REGION Network 5: RIO02 4P, 4S Vent A and Vent B control
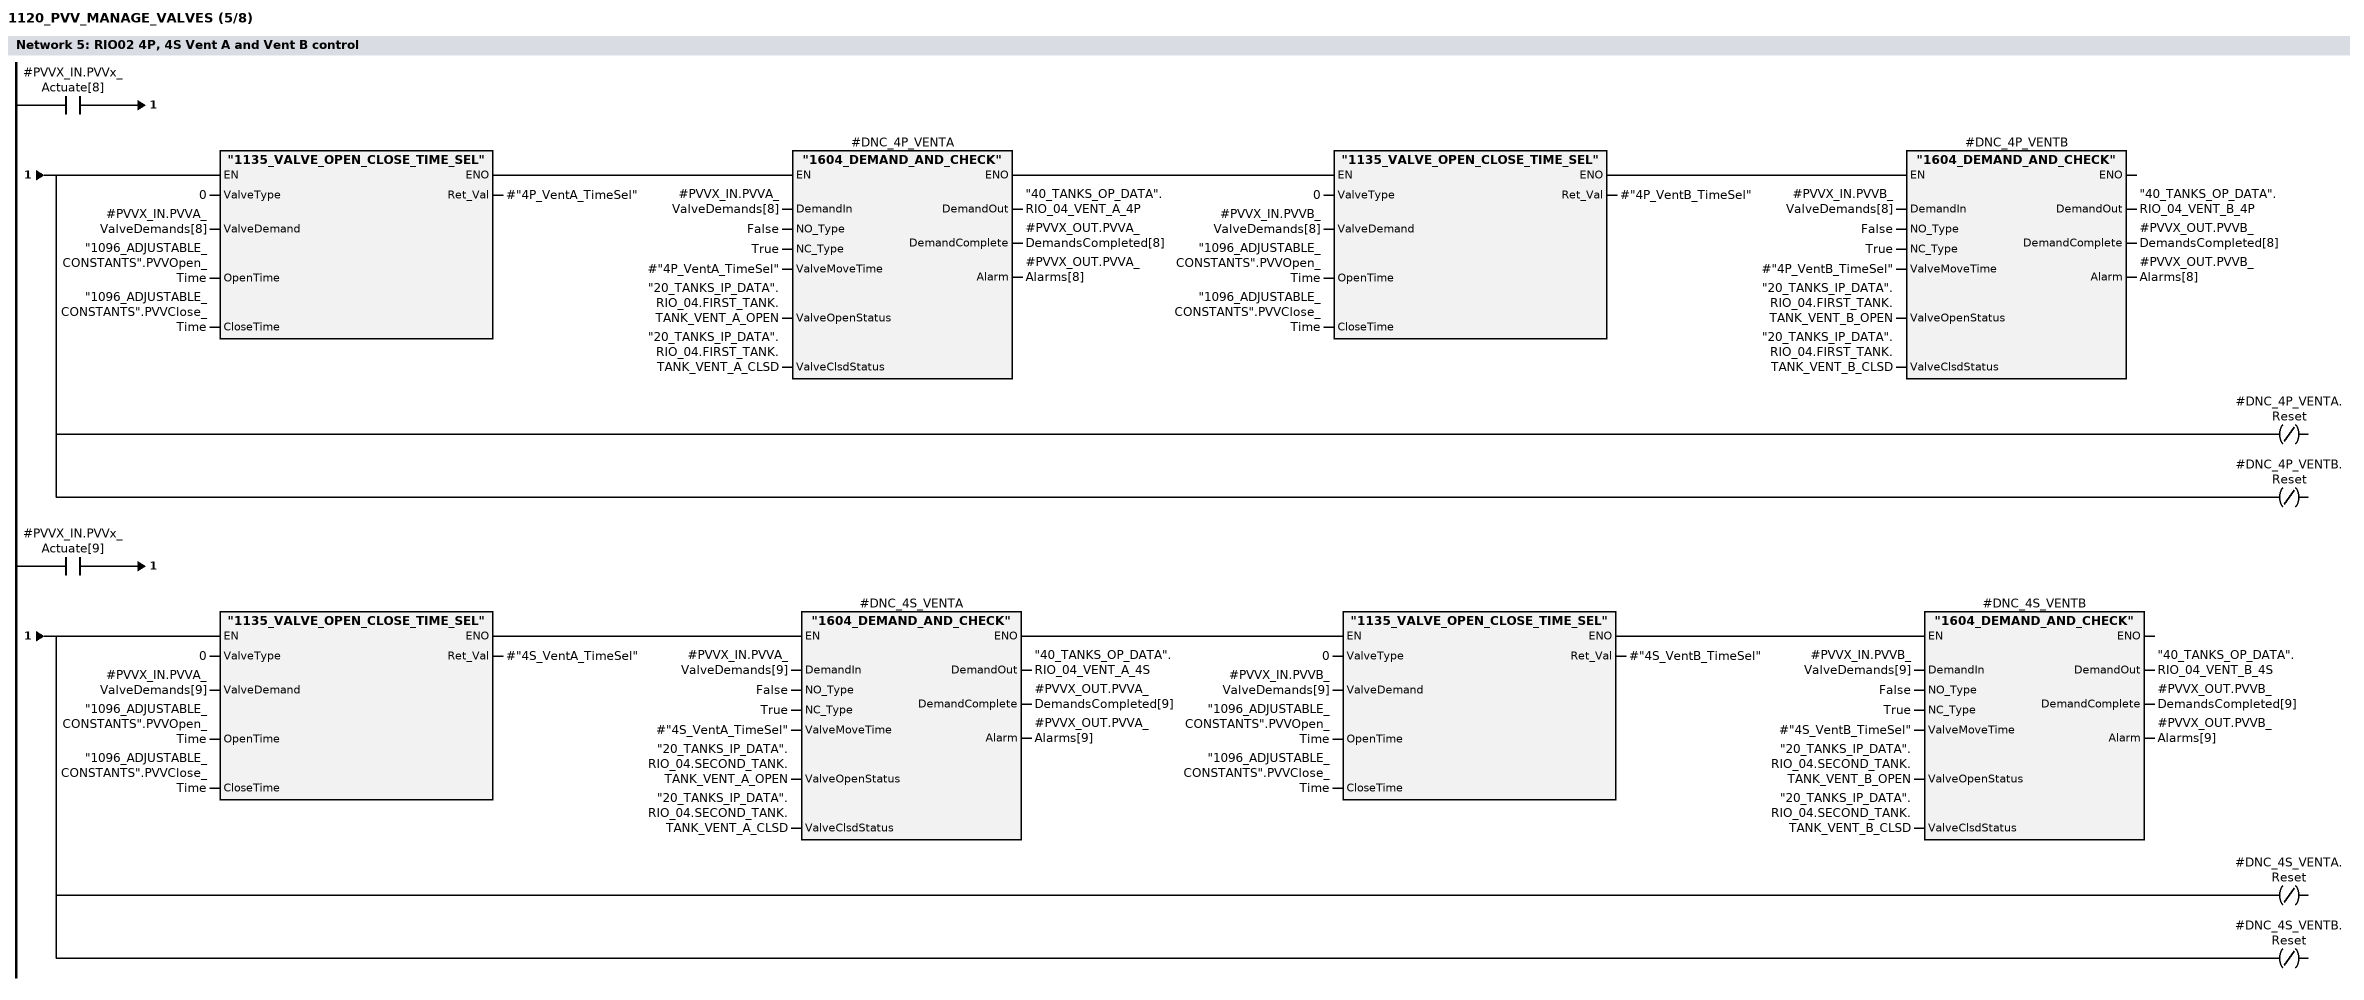
   RUNG wire#powerrail
      Contact( #PVVX_IN.PVVx_Actuate[8] )
      wire#w1
      "1135_VALVE_OPEN_CLOSE_TIME_SEL"(ValveType := 0, ValveDemand := #PVVX_IN.PVVA_ValveDemands[8], OpenTime := "1096_ADJUSTABLE_CONSTANTS".PVVOpen_Time, CloseTime := "1096_ADJUSTABLE_CONSTANTS".PVVClose_Time, Ret_Val => #"4P_VentA_TimeSel")
      #DNC_4P_VENTA(DemandIn := #PVVX_IN.PVVA_ValveDemands[8], NO_Type := False, NC_Type := True, ValveMoveTime := #"4P_VentA_TimeSel", ValveOpenStatus := "20_TANKS_IP_DATA".RIO_04.FIRST_TANK.TANK_VENT_A_OPEN, ValveClsdStatus := "20_TANKS_IP_DATA".RIO_04.FIRST_TANK.TANK_VENT_A_CLSD, DemandOut => "40_TANKS_OP_DATA".RIO_04_VENT_A_4P, DemandComplete => #PVVX_OUT.PVVA_DemandsCompleted[8], Alarm => #PVVX_OUT.PVVA_Alarms[8])
      "1135_VALVE_OPEN_CLOSE_TIME_SEL"(ValveType := 0, ValveDemand := #PVVX_IN.PVVB_ValveDemands[8], OpenTime := "1096_ADJUSTABLE_CONSTANTS".PVVOpen_Time, CloseTime := "1096_ADJUSTABLE_CONSTANTS".PVVClose_Time, Ret_Val => #"4P_VentB_TimeSel")
      #DNC_4P_VENTB(DemandIn := #PVVX_IN.PVVB_ValveDemands[8], NO_Type := False, NC_Type := True, ValveMoveTime := #"4P_VentB_TimeSel", ValveOpenStatus := "20_TANKS_IP_DATA".RIO_04.FIRST_TANK.TANK_VENT_B_OPEN, ValveClsdStatus := "20_TANKS_IP_DATA".RIO_04.FIRST_TANK.TANK_VENT_B_CLSD, DemandOut => "40_TANKS_OP_DATA".RIO_04_VENT_B_4P, DemandComplete => #PVVX_OUT.PVVB_DemandsCompleted[8], Alarm => #PVVX_OUT.PVVB_Alarms[8])
   END_RUNG
   RUNG wire#w1
      I_Coil( #DNC_4P_VENTA.Reset )
   END_RUNG
   RUNG wire#w1
      I_Coil( #DNC_4P_VENTB.Reset )
   END_RUNG
   RUNG wire#powerrail
      Contact( #PVVX_IN.PVVx_Actuate[9] )
      wire#w2
      "1135_VALVE_OPEN_CLOSE_TIME_SEL"(ValveType := 0, ValveDemand := #PVVX_IN.PVVA_ValveDemands[9], OpenTime := "1096_ADJUSTABLE_CONSTANTS".PVVOpen_Time, CloseTime := "1096_ADJUSTABLE_CONSTANTS".PVVClose_Time, Ret_Val => #"4S_VentA_TimeSel")
      #DNC_4S_VENTA(DemandIn := #PVVX_IN.PVVA_ValveDemands[9], NO_Type := False, NC_Type := True, ValveMoveTime := #"4S_VentA_TimeSel", ValveOpenStatus := "20_TANKS_IP_DATA".RIO_04.SECOND_TANK.TANK_VENT_A_OPEN, ValveClsdStatus := "20_TANKS_IP_DATA".RIO_04.SECOND_TANK.TANK_VENT_A_CLSD, DemandOut => "40_TANKS_OP_DATA".RIO_04_VENT_A_4S, DemandComplete => #PVVX_OUT.PVVA_DemandsCompleted[9], Alarm => #PVVX_OUT.PVVA_Alarms[9])
      "1135_VALVE_OPEN_CLOSE_TIME_SEL"(ValveType := 0, ValveDemand := #PVVX_IN.PVVB_ValveDemands[9], OpenTime := "1096_ADJUSTABLE_CONSTANTS".PVVOpen_Time, CloseTime := "1096_ADJUSTABLE_CONSTANTS".PVVClose_Time, Ret_Val => #"4S_VentB_TimeSel")
      #DNC_4S_VENTB(DemandIn := #PVVX_IN.PVVB_ValveDemands[9], NO_Type := False, NC_Type := True, ValveMoveTime := #"4S_VentB_TimeSel", ValveOpenStatus := "20_TANKS_IP_DATA".RIO_04.SECOND_TANK.TANK_VENT_B_OPEN, ValveClsdStatus := "20_TANKS_IP_DATA".RIO_04.SECOND_TANK.TANK_VENT_B_CLSD, DemandOut => "40_TANKS_OP_DATA".RIO_04_VENT_B_4S, DemandComplete => #PVVX_OUT.PVVB_DemandsCompleted[9], Alarm => #PVVX_OUT.PVVB_Alarms[9])
   END_RUNG
   RUNG wire#w2
      I_Coil( #DNC_4S_VENTA.Reset )
   END_RUNG
   RUNG wire#w2
      I_Coil( #DNC_4S_VENTB.Reset )
   END_RUNG
   // the same network as SCL:
   #"4P_VentA_TimeSel" := "1135_VALVE_OPEN_CLOSE_TIME_SEL"(EN := #PVVX_IN.PVVx_Actuate[8],
                           ValveType := 0,
                           ValveDemand := #PVVX_IN.PVVA_ValveDemands[8],
                           OpenTime := "1096_ADJUSTABLE_CONSTANTS".PVVOpen_Time,
                           CloseTime := "1096_ADJUSTABLE_CONSTANTS".PVVClose_Time,
                           ENO => #_w1);
   #DNC_4P_VENTA(EN := #_w1,   // "1604_DEMAND_AND_CHECK"
                 DemandIn := #PVVX_IN.PVVA_ValveDemands[8],
                 NO_Type := False,
                 NC_Type := True,
                 ValveMoveTime := #"4P_VentA_TimeSel",
                 ValveOpenStatus := "20_TANKS_IP_DATA".RIO_04.FIRST_TANK.TANK_VENT_A_OPEN,
                 ValveClsdStatus := "20_TANKS_IP_DATA".RIO_04.FIRST_TANK.TANK_VENT_A_CLSD,
                 DemandOut => "40_TANKS_OP_DATA".RIO_04_VENT_A_4P,
                 DemandComplete => #PVVX_OUT.PVVA_DemandsCompleted[8],
                 Alarm => #PVVX_OUT.PVVA_Alarms[8],
                 ENO => #_w2);
   #"4P_VentB_TimeSel" := "1135_VALVE_OPEN_CLOSE_TIME_SEL"(EN := #_w2,
                           ValveType := 0,
                           ValveDemand := #PVVX_IN.PVVB_ValveDemands[8],
                           OpenTime := "1096_ADJUSTABLE_CONSTANTS".PVVOpen_Time,
                           CloseTime := "1096_ADJUSTABLE_CONSTANTS".PVVClose_Time,
                           ENO => #_w3);
   IF #_w3 THEN
       #DNC_4P_VENTB(DemandIn := #PVVX_IN.PVVB_ValveDemands[8],   // "1604_DEMAND_AND_CHECK"
                     NO_Type := False,
                     NC_Type := True,
                     ValveMoveTime := #"4P_VentB_TimeSel",
                     ValveOpenStatus := "20_TANKS_IP_DATA".RIO_04.FIRST_TANK.TANK_VENT_B_OPEN,
                     ValveClsdStatus := "20_TANKS_IP_DATA".RIO_04.FIRST_TANK.TANK_VENT_B_CLSD,
                     DemandOut => "40_TANKS_OP_DATA".RIO_04_VENT_B_4P,
                     DemandComplete => #PVVX_OUT.PVVB_DemandsCompleted[8],
                     Alarm => #PVVX_OUT.PVVB_Alarms[8]);
   END_IF;
   #DNC_4P_VENTA.Reset := NOT #PVVX_IN.PVVx_Actuate[8];
   #DNC_4P_VENTB.Reset := NOT #PVVX_IN.PVVx_Actuate[8];
   #"4S_VentA_TimeSel" := "1135_VALVE_OPEN_CLOSE_TIME_SEL"(EN := #PVVX_IN.PVVx_Actuate[9],
                           ValveType := 0,
                           ValveDemand := #PVVX_IN.PVVA_ValveDemands[9],
                           OpenTime := "1096_ADJUSTABLE_CONSTANTS".PVVOpen_Time,
                           CloseTime := "1096_ADJUSTABLE_CONSTANTS".PVVClose_Time,
                           ENO => #_w4);
   #DNC_4S_VENTA(EN := #_w4,   // "1604_DEMAND_AND_CHECK"
                 DemandIn := #PVVX_IN.PVVA_ValveDemands[9],
                 NO_Type := False,
                 NC_Type := True,
                 ValveMoveTime := #"4S_VentA_TimeSel",
                 ValveOpenStatus := "20_TANKS_IP_DATA".RIO_04.SECOND_TANK.TANK_VENT_A_OPEN,
                 ValveClsdStatus := "20_TANKS_IP_DATA".RIO_04.SECOND_TANK.TANK_VENT_A_CLSD,
                 DemandOut => "40_TANKS_OP_DATA".RIO_04_VENT_A_4S,
                 DemandComplete => #PVVX_OUT.PVVA_DemandsCompleted[9],
                 Alarm => #PVVX_OUT.PVVA_Alarms[9],
                 ENO => #_w5);
   #"4S_VentB_TimeSel" := "1135_VALVE_OPEN_CLOSE_TIME_SEL"(EN := #_w5,
                           ValveType := 0,
                           ValveDemand := #PVVX_IN.PVVB_ValveDemands[9],
                           OpenTime := "1096_ADJUSTABLE_CONSTANTS".PVVOpen_Time,
                           CloseTime := "1096_ADJUSTABLE_CONSTANTS".PVVClose_Time,
                           ENO => #_w6);
   IF #_w6 THEN
       #DNC_4S_VENTB(DemandIn := #PVVX_IN.PVVB_ValveDemands[9],   // "1604_DEMAND_AND_CHECK"
                     NO_Type := False,
                     NC_Type := True,
                     ValveMoveTime := #"4S_VentB_TimeSel",
                     ValveOpenStatus := "20_TANKS_IP_DATA".RIO_04.SECOND_TANK.TANK_VENT_B_OPEN,
                     ValveClsdStatus := "20_TANKS_IP_DATA".RIO_04.SECOND_TANK.TANK_VENT_B_CLSD,
                     DemandOut => "40_TANKS_OP_DATA".RIO_04_VENT_B_4S,
                     DemandComplete => #PVVX_OUT.PVVB_DemandsCompleted[9],
                     Alarm => #PVVX_OUT.PVVB_Alarms[9]);
   END_IF;
   #DNC_4S_VENTA.Reset := NOT #PVVX_IN.PVVx_Actuate[9];
   #DNC_4S_VENTB.Reset := NOT #PVVX_IN.PVVx_Actuate[9];
END_REGION

REGION Network 6: RIO02 5P, 5S Vent A and Vent B control
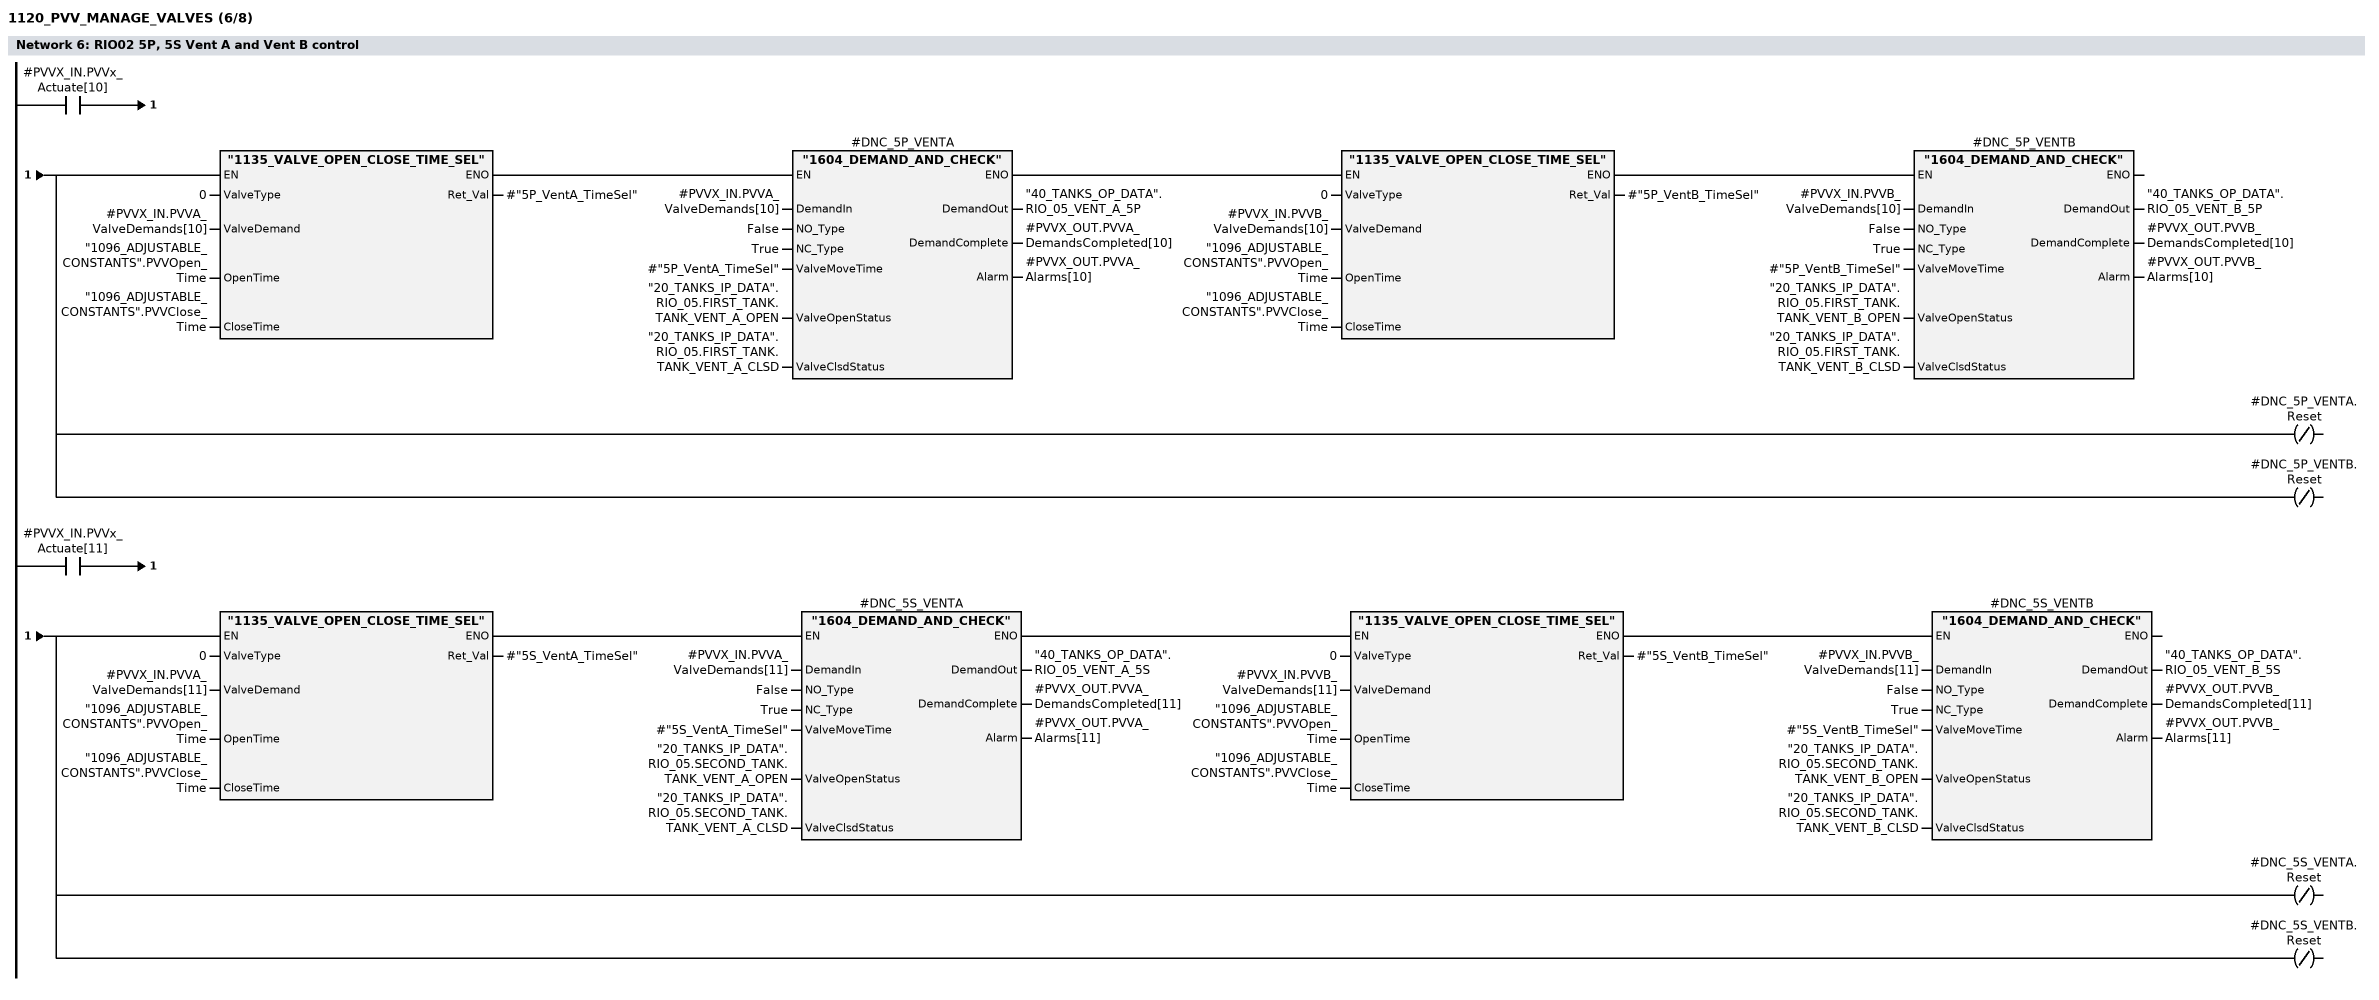
   RUNG wire#powerrail
      Contact( #PVVX_IN.PVVx_Actuate[10] )
      wire#w1
      "1135_VALVE_OPEN_CLOSE_TIME_SEL"(ValveType := 0, ValveDemand := #PVVX_IN.PVVA_ValveDemands[10], OpenTime := "1096_ADJUSTABLE_CONSTANTS".PVVOpen_Time, CloseTime := "1096_ADJUSTABLE_CONSTANTS".PVVClose_Time, Ret_Val => #"5P_VentA_TimeSel")
      #DNC_5P_VENTA(DemandIn := #PVVX_IN.PVVA_ValveDemands[10], NO_Type := False, NC_Type := True, ValveMoveTime := #"5P_VentA_TimeSel", ValveOpenStatus := "20_TANKS_IP_DATA".RIO_05.FIRST_TANK.TANK_VENT_A_OPEN, ValveClsdStatus := "20_TANKS_IP_DATA".RIO_05.FIRST_TANK.TANK_VENT_A_CLSD, DemandOut => "40_TANKS_OP_DATA".RIO_05_VENT_A_5P, DemandComplete => #PVVX_OUT.PVVA_DemandsCompleted[10], Alarm => #PVVX_OUT.PVVA_Alarms[10])
      "1135_VALVE_OPEN_CLOSE_TIME_SEL"(ValveType := 0, ValveDemand := #PVVX_IN.PVVB_ValveDemands[10], OpenTime := "1096_ADJUSTABLE_CONSTANTS".PVVOpen_Time, CloseTime := "1096_ADJUSTABLE_CONSTANTS".PVVClose_Time, Ret_Val => #"5P_VentB_TimeSel")
      #DNC_5P_VENTB(DemandIn := #PVVX_IN.PVVB_ValveDemands[10], NO_Type := False, NC_Type := True, ValveMoveTime := #"5P_VentB_TimeSel", ValveOpenStatus := "20_TANKS_IP_DATA".RIO_05.FIRST_TANK.TANK_VENT_B_OPEN, ValveClsdStatus := "20_TANKS_IP_DATA".RIO_05.FIRST_TANK.TANK_VENT_B_CLSD, DemandOut => "40_TANKS_OP_DATA".RIO_05_VENT_B_5P, DemandComplete => #PVVX_OUT.PVVB_DemandsCompleted[10], Alarm => #PVVX_OUT.PVVB_Alarms[10])
   END_RUNG
   RUNG wire#w1
      I_Coil( #DNC_5P_VENTA.Reset )
   END_RUNG
   RUNG wire#w1
      I_Coil( #DNC_5P_VENTB.Reset )
   END_RUNG
   RUNG wire#powerrail
      Contact( #PVVX_IN.PVVx_Actuate[11] )
      wire#w2
      "1135_VALVE_OPEN_CLOSE_TIME_SEL"(ValveType := 0, ValveDemand := #PVVX_IN.PVVA_ValveDemands[11], OpenTime := "1096_ADJUSTABLE_CONSTANTS".PVVOpen_Time, CloseTime := "1096_ADJUSTABLE_CONSTANTS".PVVClose_Time, Ret_Val => #"5S_VentA_TimeSel")
      #DNC_5S_VENTA(DemandIn := #PVVX_IN.PVVA_ValveDemands[11], NO_Type := False, NC_Type := True, ValveMoveTime := #"5S_VentA_TimeSel", ValveOpenStatus := "20_TANKS_IP_DATA".RIO_05.SECOND_TANK.TANK_VENT_A_OPEN, ValveClsdStatus := "20_TANKS_IP_DATA".RIO_05.SECOND_TANK.TANK_VENT_A_CLSD, DemandOut => "40_TANKS_OP_DATA".RIO_05_VENT_A_5S, DemandComplete => #PVVX_OUT.PVVA_DemandsCompleted[11], Alarm => #PVVX_OUT.PVVA_Alarms[11])
      "1135_VALVE_OPEN_CLOSE_TIME_SEL"(ValveType := 0, ValveDemand := #PVVX_IN.PVVB_ValveDemands[11], OpenTime := "1096_ADJUSTABLE_CONSTANTS".PVVOpen_Time, CloseTime := "1096_ADJUSTABLE_CONSTANTS".PVVClose_Time, Ret_Val => #"5S_VentB_TimeSel")
      #DNC_5S_VENTB(DemandIn := #PVVX_IN.PVVB_ValveDemands[11], NO_Type := False, NC_Type := True, ValveMoveTime := #"5S_VentB_TimeSel", ValveOpenStatus := "20_TANKS_IP_DATA".RIO_05.SECOND_TANK.TANK_VENT_B_OPEN, ValveClsdStatus := "20_TANKS_IP_DATA".RIO_05.SECOND_TANK.TANK_VENT_B_CLSD, DemandOut => "40_TANKS_OP_DATA".RIO_05_VENT_B_5S, DemandComplete => #PVVX_OUT.PVVB_DemandsCompleted[11], Alarm => #PVVX_OUT.PVVB_Alarms[11])
   END_RUNG
   RUNG wire#w2
      I_Coil( #DNC_5S_VENTA.Reset )
   END_RUNG
   RUNG wire#w2
      I_Coil( #DNC_5S_VENTB.Reset )
   END_RUNG
   // the same network as SCL:
   #"5P_VentA_TimeSel" := "1135_VALVE_OPEN_CLOSE_TIME_SEL"(EN := #PVVX_IN.PVVx_Actuate[10],
                           ValveType := 0,
                           ValveDemand := #PVVX_IN.PVVA_ValveDemands[10],
                           OpenTime := "1096_ADJUSTABLE_CONSTANTS".PVVOpen_Time,
                           CloseTime := "1096_ADJUSTABLE_CONSTANTS".PVVClose_Time,
                           ENO => #_w1);
   #DNC_5P_VENTA(EN := #_w1,   // "1604_DEMAND_AND_CHECK"
                 DemandIn := #PVVX_IN.PVVA_ValveDemands[10],
                 NO_Type := False,
                 NC_Type := True,
                 ValveMoveTime := #"5P_VentA_TimeSel",
                 ValveOpenStatus := "20_TANKS_IP_DATA".RIO_05.FIRST_TANK.TANK_VENT_A_OPEN,
                 ValveClsdStatus := "20_TANKS_IP_DATA".RIO_05.FIRST_TANK.TANK_VENT_A_CLSD,
                 DemandOut => "40_TANKS_OP_DATA".RIO_05_VENT_A_5P,
                 DemandComplete => #PVVX_OUT.PVVA_DemandsCompleted[10],
                 Alarm => #PVVX_OUT.PVVA_Alarms[10],
                 ENO => #_w2);
   #"5P_VentB_TimeSel" := "1135_VALVE_OPEN_CLOSE_TIME_SEL"(EN := #_w2,
                           ValveType := 0,
                           ValveDemand := #PVVX_IN.PVVB_ValveDemands[10],
                           OpenTime := "1096_ADJUSTABLE_CONSTANTS".PVVOpen_Time,
                           CloseTime := "1096_ADJUSTABLE_CONSTANTS".PVVClose_Time,
                           ENO => #_w3);
   IF #_w3 THEN
       #DNC_5P_VENTB(DemandIn := #PVVX_IN.PVVB_ValveDemands[10],   // "1604_DEMAND_AND_CHECK"
                     NO_Type := False,
                     NC_Type := True,
                     ValveMoveTime := #"5P_VentB_TimeSel",
                     ValveOpenStatus := "20_TANKS_IP_DATA".RIO_05.FIRST_TANK.TANK_VENT_B_OPEN,
                     ValveClsdStatus := "20_TANKS_IP_DATA".RIO_05.FIRST_TANK.TANK_VENT_B_CLSD,
                     DemandOut => "40_TANKS_OP_DATA".RIO_05_VENT_B_5P,
                     DemandComplete => #PVVX_OUT.PVVB_DemandsCompleted[10],
                     Alarm => #PVVX_OUT.PVVB_Alarms[10]);
   END_IF;
   #DNC_5P_VENTA.Reset := NOT #PVVX_IN.PVVx_Actuate[10];
   #DNC_5P_VENTB.Reset := NOT #PVVX_IN.PVVx_Actuate[10];
   #"5S_VentA_TimeSel" := "1135_VALVE_OPEN_CLOSE_TIME_SEL"(EN := #PVVX_IN.PVVx_Actuate[11],
                           ValveType := 0,
                           ValveDemand := #PVVX_IN.PVVA_ValveDemands[11],
                           OpenTime := "1096_ADJUSTABLE_CONSTANTS".PVVOpen_Time,
                           CloseTime := "1096_ADJUSTABLE_CONSTANTS".PVVClose_Time,
                           ENO => #_w4);
   #DNC_5S_VENTA(EN := #_w4,   // "1604_DEMAND_AND_CHECK"
                 DemandIn := #PVVX_IN.PVVA_ValveDemands[11],
                 NO_Type := False,
                 NC_Type := True,
                 ValveMoveTime := #"5S_VentA_TimeSel",
                 ValveOpenStatus := "20_TANKS_IP_DATA".RIO_05.SECOND_TANK.TANK_VENT_A_OPEN,
                 ValveClsdStatus := "20_TANKS_IP_DATA".RIO_05.SECOND_TANK.TANK_VENT_A_CLSD,
                 DemandOut => "40_TANKS_OP_DATA".RIO_05_VENT_A_5S,
                 DemandComplete => #PVVX_OUT.PVVA_DemandsCompleted[11],
                 Alarm => #PVVX_OUT.PVVA_Alarms[11],
                 ENO => #_w5);
   #"5S_VentB_TimeSel" := "1135_VALVE_OPEN_CLOSE_TIME_SEL"(EN := #_w5,
                           ValveType := 0,
                           ValveDemand := #PVVX_IN.PVVB_ValveDemands[11],
                           OpenTime := "1096_ADJUSTABLE_CONSTANTS".PVVOpen_Time,
                           CloseTime := "1096_ADJUSTABLE_CONSTANTS".PVVClose_Time,
                           ENO => #_w6);
   IF #_w6 THEN
       #DNC_5S_VENTB(DemandIn := #PVVX_IN.PVVB_ValveDemands[11],   // "1604_DEMAND_AND_CHECK"
                     NO_Type := False,
                     NC_Type := True,
                     ValveMoveTime := #"5S_VentB_TimeSel",
                     ValveOpenStatus := "20_TANKS_IP_DATA".RIO_05.SECOND_TANK.TANK_VENT_B_OPEN,
                     ValveClsdStatus := "20_TANKS_IP_DATA".RIO_05.SECOND_TANK.TANK_VENT_B_CLSD,
                     DemandOut => "40_TANKS_OP_DATA".RIO_05_VENT_B_5S,
                     DemandComplete => #PVVX_OUT.PVVB_DemandsCompleted[11],
                     Alarm => #PVVX_OUT.PVVB_Alarms[11]);
   END_IF;
   #DNC_5S_VENTA.Reset := NOT #PVVX_IN.PVVx_Actuate[11];
   #DNC_5S_VENTB.Reset := NOT #PVVX_IN.PVVx_Actuate[11];
END_REGION

REGION Network 7: RIO02 6P, 6S Vent A and Vent B control
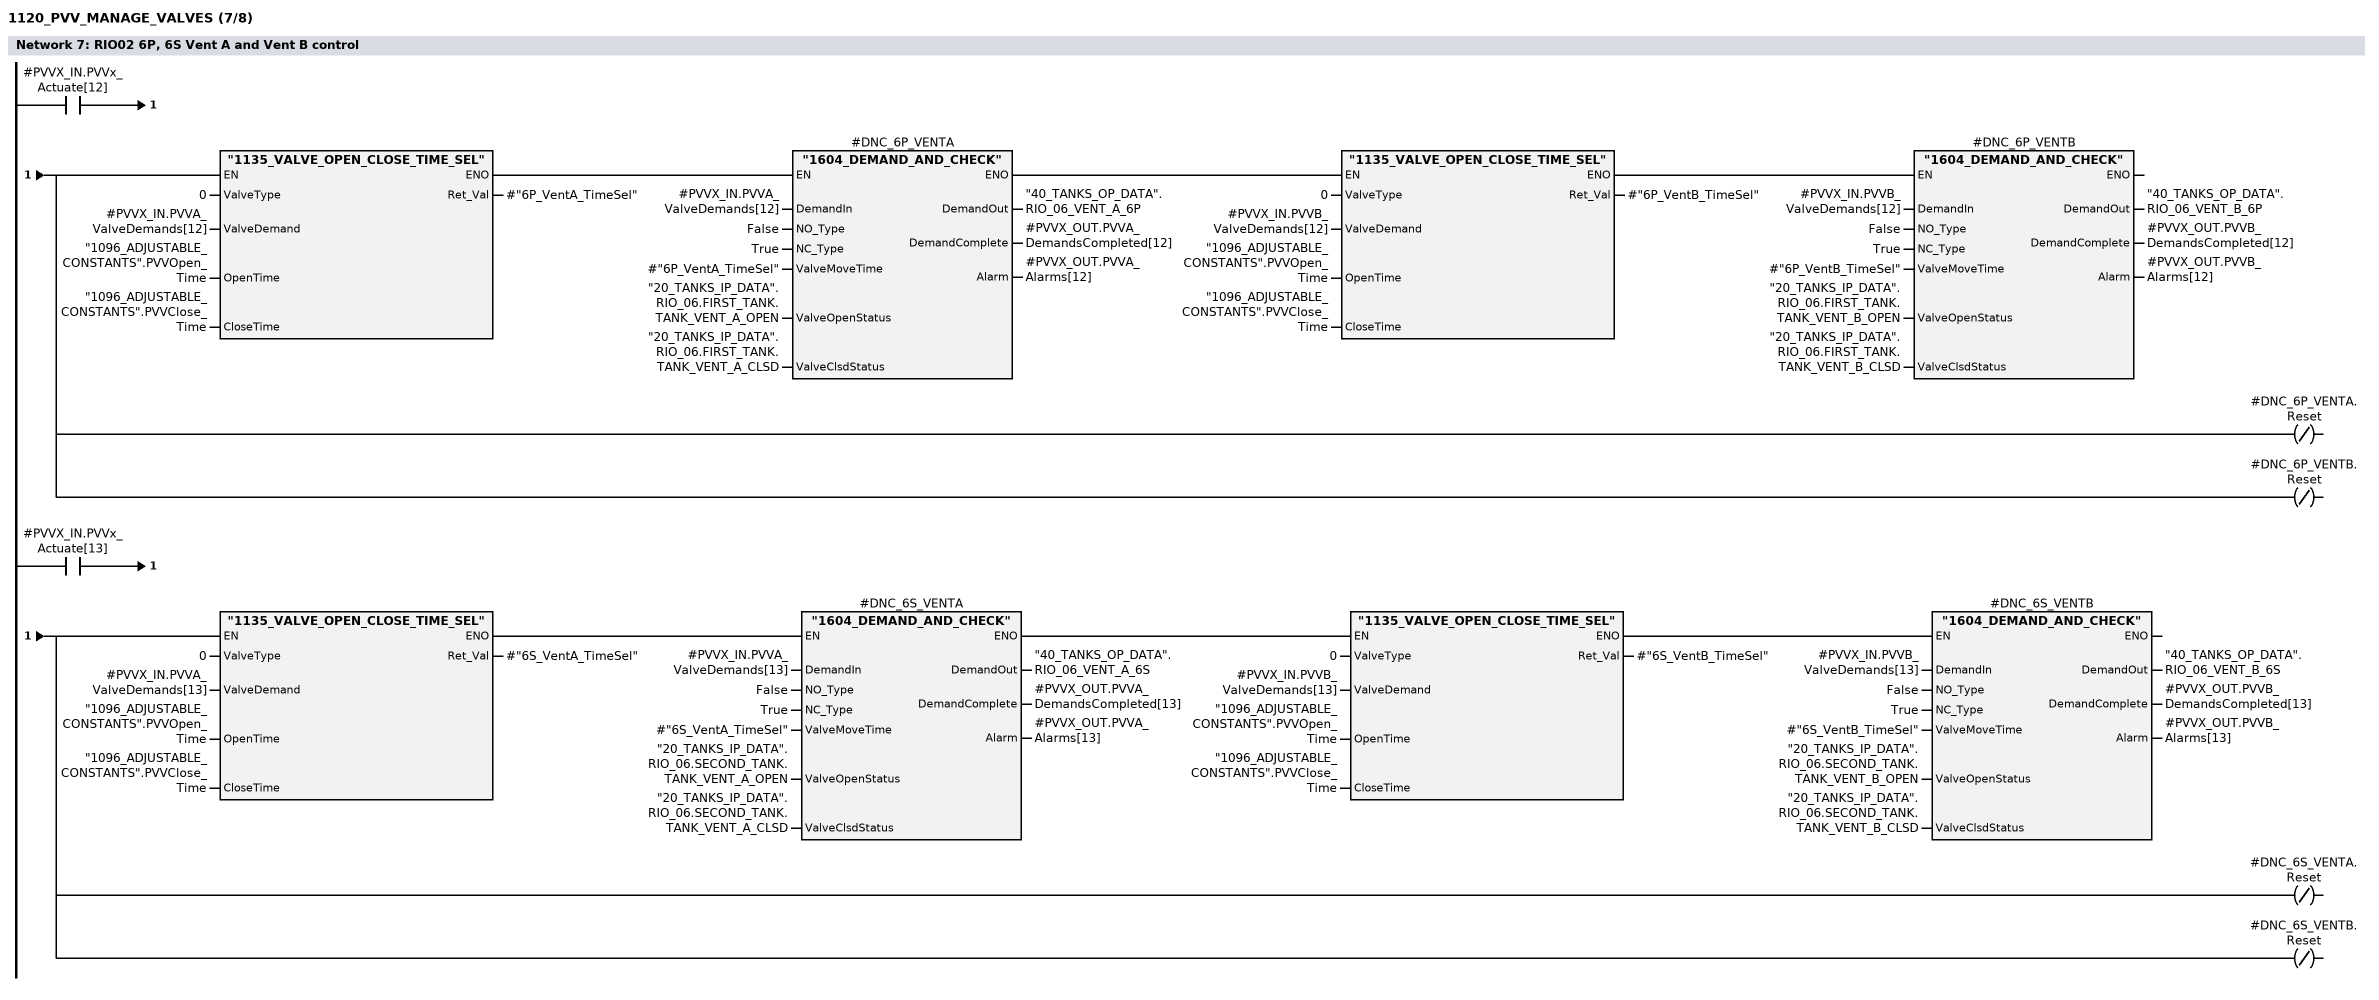
   RUNG wire#powerrail
      Contact( #PVVX_IN.PVVx_Actuate[12] )
      wire#w1
      "1135_VALVE_OPEN_CLOSE_TIME_SEL"(ValveType := 0, ValveDemand := #PVVX_IN.PVVA_ValveDemands[12], OpenTime := "1096_ADJUSTABLE_CONSTANTS".PVVOpen_Time, CloseTime := "1096_ADJUSTABLE_CONSTANTS".PVVClose_Time, Ret_Val => #"6P_VentA_TimeSel")
      #DNC_6P_VENTA(DemandIn := #PVVX_IN.PVVA_ValveDemands[12], NO_Type := False, NC_Type := True, ValveMoveTime := #"6P_VentA_TimeSel", ValveOpenStatus := "20_TANKS_IP_DATA".RIO_06.FIRST_TANK.TANK_VENT_A_OPEN, ValveClsdStatus := "20_TANKS_IP_DATA".RIO_06.FIRST_TANK.TANK_VENT_A_CLSD, DemandOut => "40_TANKS_OP_DATA".RIO_06_VENT_A_6P, DemandComplete => #PVVX_OUT.PVVA_DemandsCompleted[12], Alarm => #PVVX_OUT.PVVA_Alarms[12])
      "1135_VALVE_OPEN_CLOSE_TIME_SEL"(ValveType := 0, ValveDemand := #PVVX_IN.PVVB_ValveDemands[12], OpenTime := "1096_ADJUSTABLE_CONSTANTS".PVVOpen_Time, CloseTime := "1096_ADJUSTABLE_CONSTANTS".PVVClose_Time, Ret_Val => #"6P_VentB_TimeSel")
      #DNC_6P_VENTB(DemandIn := #PVVX_IN.PVVB_ValveDemands[12], NO_Type := False, NC_Type := True, ValveMoveTime := #"6P_VentB_TimeSel", ValveOpenStatus := "20_TANKS_IP_DATA".RIO_06.FIRST_TANK.TANK_VENT_B_OPEN, ValveClsdStatus := "20_TANKS_IP_DATA".RIO_06.FIRST_TANK.TANK_VENT_B_CLSD, DemandOut => "40_TANKS_OP_DATA".RIO_06_VENT_B_6P, DemandComplete => #PVVX_OUT.PVVB_DemandsCompleted[12], Alarm => #PVVX_OUT.PVVB_Alarms[12])
   END_RUNG
   RUNG wire#w1
      I_Coil( #DNC_6P_VENTA.Reset )
   END_RUNG
   RUNG wire#w1
      I_Coil( #DNC_6P_VENTB.Reset )
   END_RUNG
   RUNG wire#powerrail
      Contact( #PVVX_IN.PVVx_Actuate[13] )
      wire#w2
      "1135_VALVE_OPEN_CLOSE_TIME_SEL"(ValveType := 0, ValveDemand := #PVVX_IN.PVVA_ValveDemands[13], OpenTime := "1096_ADJUSTABLE_CONSTANTS".PVVOpen_Time, CloseTime := "1096_ADJUSTABLE_CONSTANTS".PVVClose_Time, Ret_Val => #"6S_VentA_TimeSel")
      #DNC_6S_VENTA(DemandIn := #PVVX_IN.PVVA_ValveDemands[13], NO_Type := False, NC_Type := True, ValveMoveTime := #"6S_VentA_TimeSel", ValveOpenStatus := "20_TANKS_IP_DATA".RIO_06.SECOND_TANK.TANK_VENT_A_OPEN, ValveClsdStatus := "20_TANKS_IP_DATA".RIO_06.SECOND_TANK.TANK_VENT_A_CLSD, DemandOut => "40_TANKS_OP_DATA".RIO_06_VENT_A_6S, DemandComplete => #PVVX_OUT.PVVA_DemandsCompleted[13], Alarm => #PVVX_OUT.PVVA_Alarms[13])
      "1135_VALVE_OPEN_CLOSE_TIME_SEL"(ValveType := 0, ValveDemand := #PVVX_IN.PVVB_ValveDemands[13], OpenTime := "1096_ADJUSTABLE_CONSTANTS".PVVOpen_Time, CloseTime := "1096_ADJUSTABLE_CONSTANTS".PVVClose_Time, Ret_Val => #"6S_VentB_TimeSel")
      #DNC_6S_VENTB(DemandIn := #PVVX_IN.PVVB_ValveDemands[13], NO_Type := False, NC_Type := True, ValveMoveTime := #"6S_VentB_TimeSel", ValveOpenStatus := "20_TANKS_IP_DATA".RIO_06.SECOND_TANK.TANK_VENT_B_OPEN, ValveClsdStatus := "20_TANKS_IP_DATA".RIO_06.SECOND_TANK.TANK_VENT_B_CLSD, DemandOut => "40_TANKS_OP_DATA".RIO_06_VENT_B_6S, DemandComplete => #PVVX_OUT.PVVB_DemandsCompleted[13], Alarm => #PVVX_OUT.PVVB_Alarms[13])
   END_RUNG
   RUNG wire#w2
      I_Coil( #DNC_6S_VENTA.Reset )
   END_RUNG
   RUNG wire#w2
      I_Coil( #DNC_6S_VENTB.Reset )
   END_RUNG
   // the same network as SCL:
   #"6P_VentA_TimeSel" := "1135_VALVE_OPEN_CLOSE_TIME_SEL"(EN := #PVVX_IN.PVVx_Actuate[12],
                           ValveType := 0,
                           ValveDemand := #PVVX_IN.PVVA_ValveDemands[12],
                           OpenTime := "1096_ADJUSTABLE_CONSTANTS".PVVOpen_Time,
                           CloseTime := "1096_ADJUSTABLE_CONSTANTS".PVVClose_Time,
                           ENO => #_w1);
   #DNC_6P_VENTA(EN := #_w1,   // "1604_DEMAND_AND_CHECK"
                 DemandIn := #PVVX_IN.PVVA_ValveDemands[12],
                 NO_Type := False,
                 NC_Type := True,
                 ValveMoveTime := #"6P_VentA_TimeSel",
                 ValveOpenStatus := "20_TANKS_IP_DATA".RIO_06.FIRST_TANK.TANK_VENT_A_OPEN,
                 ValveClsdStatus := "20_TANKS_IP_DATA".RIO_06.FIRST_TANK.TANK_VENT_A_CLSD,
                 DemandOut => "40_TANKS_OP_DATA".RIO_06_VENT_A_6P,
                 DemandComplete => #PVVX_OUT.PVVA_DemandsCompleted[12],
                 Alarm => #PVVX_OUT.PVVA_Alarms[12],
                 ENO => #_w2);
   #"6P_VentB_TimeSel" := "1135_VALVE_OPEN_CLOSE_TIME_SEL"(EN := #_w2,
                           ValveType := 0,
                           ValveDemand := #PVVX_IN.PVVB_ValveDemands[12],
                           OpenTime := "1096_ADJUSTABLE_CONSTANTS".PVVOpen_Time,
                           CloseTime := "1096_ADJUSTABLE_CONSTANTS".PVVClose_Time,
                           ENO => #_w3);
   IF #_w3 THEN
       #DNC_6P_VENTB(DemandIn := #PVVX_IN.PVVB_ValveDemands[12],   // "1604_DEMAND_AND_CHECK"
                     NO_Type := False,
                     NC_Type := True,
                     ValveMoveTime := #"6P_VentB_TimeSel",
                     ValveOpenStatus := "20_TANKS_IP_DATA".RIO_06.FIRST_TANK.TANK_VENT_B_OPEN,
                     ValveClsdStatus := "20_TANKS_IP_DATA".RIO_06.FIRST_TANK.TANK_VENT_B_CLSD,
                     DemandOut => "40_TANKS_OP_DATA".RIO_06_VENT_B_6P,
                     DemandComplete => #PVVX_OUT.PVVB_DemandsCompleted[12],
                     Alarm => #PVVX_OUT.PVVB_Alarms[12]);
   END_IF;
   #DNC_6P_VENTA.Reset := NOT #PVVX_IN.PVVx_Actuate[12];
   #DNC_6P_VENTB.Reset := NOT #PVVX_IN.PVVx_Actuate[12];
   #"6S_VentA_TimeSel" := "1135_VALVE_OPEN_CLOSE_TIME_SEL"(EN := #PVVX_IN.PVVx_Actuate[13],
                           ValveType := 0,
                           ValveDemand := #PVVX_IN.PVVA_ValveDemands[13],
                           OpenTime := "1096_ADJUSTABLE_CONSTANTS".PVVOpen_Time,
                           CloseTime := "1096_ADJUSTABLE_CONSTANTS".PVVClose_Time,
                           ENO => #_w4);
   #DNC_6S_VENTA(EN := #_w4,   // "1604_DEMAND_AND_CHECK"
                 DemandIn := #PVVX_IN.PVVA_ValveDemands[13],
                 NO_Type := False,
                 NC_Type := True,
                 ValveMoveTime := #"6S_VentA_TimeSel",
                 ValveOpenStatus := "20_TANKS_IP_DATA".RIO_06.SECOND_TANK.TANK_VENT_A_OPEN,
                 ValveClsdStatus := "20_TANKS_IP_DATA".RIO_06.SECOND_TANK.TANK_VENT_A_CLSD,
                 DemandOut => "40_TANKS_OP_DATA".RIO_06_VENT_A_6S,
                 DemandComplete => #PVVX_OUT.PVVA_DemandsCompleted[13],
                 Alarm => #PVVX_OUT.PVVA_Alarms[13],
                 ENO => #_w5);
   #"6S_VentB_TimeSel" := "1135_VALVE_OPEN_CLOSE_TIME_SEL"(EN := #_w5,
                           ValveType := 0,
                           ValveDemand := #PVVX_IN.PVVB_ValveDemands[13],
                           OpenTime := "1096_ADJUSTABLE_CONSTANTS".PVVOpen_Time,
                           CloseTime := "1096_ADJUSTABLE_CONSTANTS".PVVClose_Time,
                           ENO => #_w6);
   IF #_w6 THEN
       #DNC_6S_VENTB(DemandIn := #PVVX_IN.PVVB_ValveDemands[13],   // "1604_DEMAND_AND_CHECK"
                     NO_Type := False,
                     NC_Type := True,
                     ValveMoveTime := #"6S_VentB_TimeSel",
                     ValveOpenStatus := "20_TANKS_IP_DATA".RIO_06.SECOND_TANK.TANK_VENT_B_OPEN,
                     ValveClsdStatus := "20_TANKS_IP_DATA".RIO_06.SECOND_TANK.TANK_VENT_B_CLSD,
                     DemandOut => "40_TANKS_OP_DATA".RIO_06_VENT_B_6S,
                     DemandComplete => #PVVX_OUT.PVVB_DemandsCompleted[13],
                     Alarm => #PVVX_OUT.PVVB_Alarms[13]);
   END_IF;
   #DNC_6S_VENTA.Reset := NOT #PVVX_IN.PVVx_Actuate[13];
   #DNC_6S_VENTB.Reset := NOT #PVVX_IN.PVVx_Actuate[13];
END_REGION

REGION Network 8: RIO07 APT Vent A and Vent B control
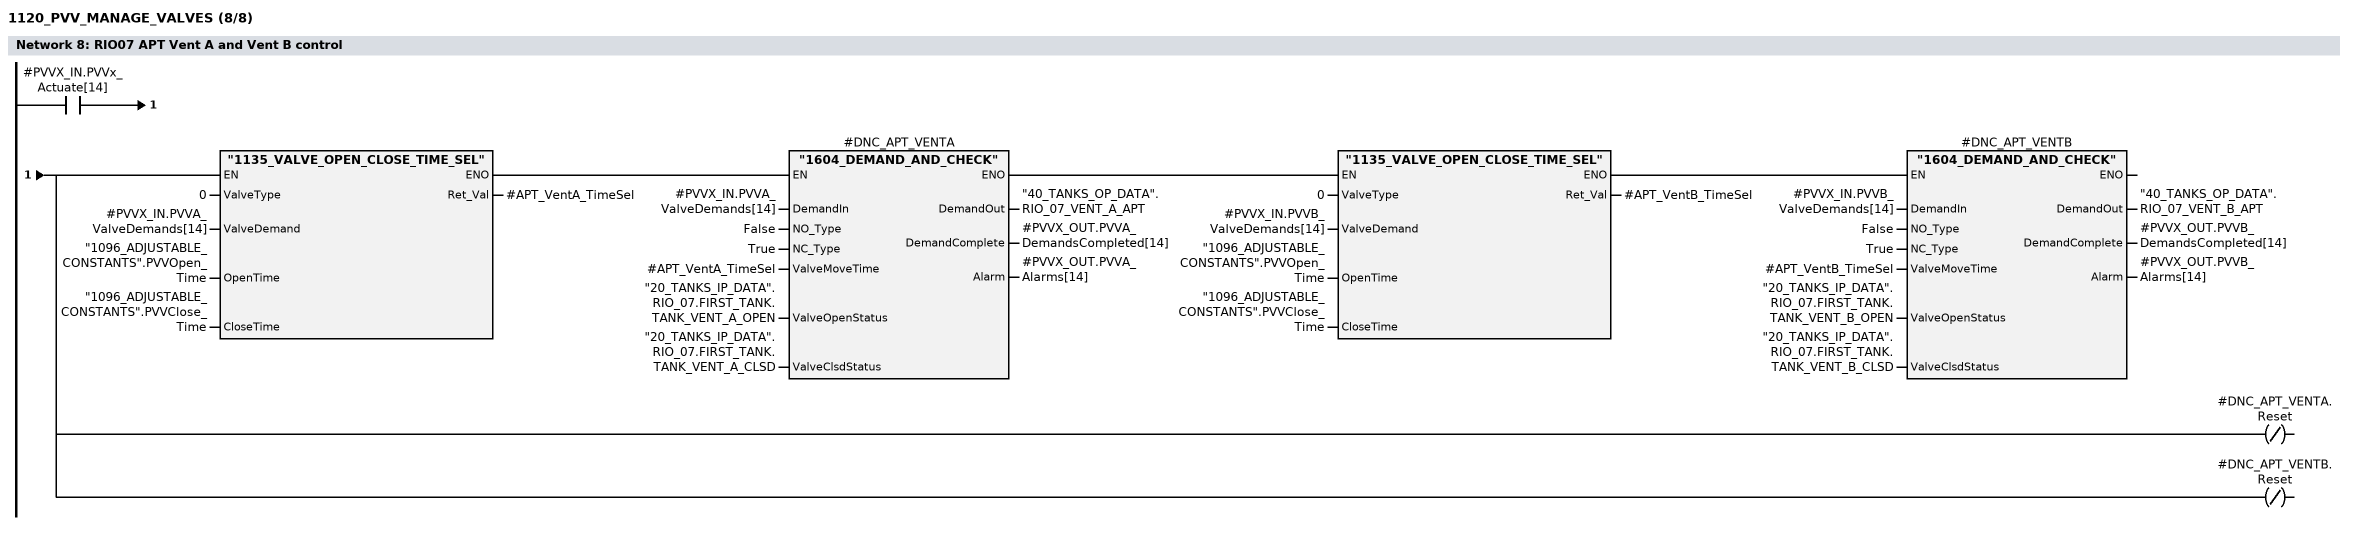
   RUNG wire#powerrail
      Contact( #PVVX_IN.PVVx_Actuate[14] )
      wire#w1
      "1135_VALVE_OPEN_CLOSE_TIME_SEL"(ValveType := 0, ValveDemand := #PVVX_IN.PVVA_ValveDemands[14], OpenTime := "1096_ADJUSTABLE_CONSTANTS".PVVOpen_Time, CloseTime := "1096_ADJUSTABLE_CONSTANTS".PVVClose_Time, Ret_Val => #APT_VentA_TimeSel)
      #DNC_APT_VENTA(DemandIn := #PVVX_IN.PVVA_ValveDemands[14], NO_Type := False, NC_Type := True, ValveMoveTime := #APT_VentA_TimeSel, ValveOpenStatus := "20_TANKS_IP_DATA".RIO_07.FIRST_TANK.TANK_VENT_A_OPEN, ValveClsdStatus := "20_TANKS_IP_DATA".RIO_07.FIRST_TANK.TANK_VENT_A_CLSD, DemandOut => "40_TANKS_OP_DATA".RIO_07_VENT_A_APT, DemandComplete => #PVVX_OUT.PVVA_DemandsCompleted[14], Alarm => #PVVX_OUT.PVVA_Alarms[14])
      "1135_VALVE_OPEN_CLOSE_TIME_SEL"(ValveType := 0, ValveDemand := #PVVX_IN.PVVB_ValveDemands[14], OpenTime := "1096_ADJUSTABLE_CONSTANTS".PVVOpen_Time, CloseTime := "1096_ADJUSTABLE_CONSTANTS".PVVClose_Time, Ret_Val => #APT_VentB_TimeSel)
      #DNC_APT_VENTB(DemandIn := #PVVX_IN.PVVB_ValveDemands[14], NO_Type := False, NC_Type := True, ValveMoveTime := #APT_VentB_TimeSel, ValveOpenStatus := "20_TANKS_IP_DATA".RIO_07.FIRST_TANK.TANK_VENT_B_OPEN, ValveClsdStatus := "20_TANKS_IP_DATA".RIO_07.FIRST_TANK.TANK_VENT_B_CLSD, DemandOut => "40_TANKS_OP_DATA".RIO_07_VENT_B_APT, DemandComplete => #PVVX_OUT.PVVB_DemandsCompleted[14], Alarm => #PVVX_OUT.PVVB_Alarms[14])
   END_RUNG
   RUNG wire#w1
      I_Coil( #DNC_APT_VENTA.Reset )
   END_RUNG
   RUNG wire#w1
      I_Coil( #DNC_APT_VENTB.Reset )
   END_RUNG
   // the same network as SCL:
   #APT_VentA_TimeSel := "1135_VALVE_OPEN_CLOSE_TIME_SEL"(EN := #PVVX_IN.PVVx_Actuate[14],
                           ValveType := 0,
                           ValveDemand := #PVVX_IN.PVVA_ValveDemands[14],
                           OpenTime := "1096_ADJUSTABLE_CONSTANTS".PVVOpen_Time,
                           CloseTime := "1096_ADJUSTABLE_CONSTANTS".PVVClose_Time,
                           ENO => #_w1);
   #DNC_APT_VENTA(EN := #_w1,   // "1604_DEMAND_AND_CHECK"
                  DemandIn := #PVVX_IN.PVVA_ValveDemands[14],
                  NO_Type := False,
                  NC_Type := True,
                  ValveMoveTime := #APT_VentA_TimeSel,
                  ValveOpenStatus := "20_TANKS_IP_DATA".RIO_07.FIRST_TANK.TANK_VENT_A_OPEN,
                  ValveClsdStatus := "20_TANKS_IP_DATA".RIO_07.FIRST_TANK.TANK_VENT_A_CLSD,
                  DemandOut => "40_TANKS_OP_DATA".RIO_07_VENT_A_APT,
                  DemandComplete => #PVVX_OUT.PVVA_DemandsCompleted[14],
                  Alarm => #PVVX_OUT.PVVA_Alarms[14],
                  ENO => #_w2);
   #APT_VentB_TimeSel := "1135_VALVE_OPEN_CLOSE_TIME_SEL"(EN := #_w2,
                           ValveType := 0,
                           ValveDemand := #PVVX_IN.PVVB_ValveDemands[14],
                           OpenTime := "1096_ADJUSTABLE_CONSTANTS".PVVOpen_Time,
                           CloseTime := "1096_ADJUSTABLE_CONSTANTS".PVVClose_Time,
                           ENO => #_w3);
   IF #_w3 THEN
       #DNC_APT_VENTB(DemandIn := #PVVX_IN.PVVB_ValveDemands[14],   // "1604_DEMAND_AND_CHECK"
                      NO_Type := False,
                      NC_Type := True,
                      ValveMoveTime := #APT_VentB_TimeSel,
                      ValveOpenStatus := "20_TANKS_IP_DATA".RIO_07.FIRST_TANK.TANK_VENT_B_OPEN,
                      ValveClsdStatus := "20_TANKS_IP_DATA".RIO_07.FIRST_TANK.TANK_VENT_B_CLSD,
                      DemandOut => "40_TANKS_OP_DATA".RIO_07_VENT_B_APT,
                      DemandComplete => #PVVX_OUT.PVVB_DemandsCompleted[14],
                      Alarm => #PVVX_OUT.PVVB_Alarms[14]);
   END_IF;
   #DNC_APT_VENTA.Reset := NOT #PVVX_IN.PVVx_Actuate[14];
   #DNC_APT_VENTB.Reset := NOT #PVVX_IN.PVVx_Actuate[14];
END_REGION
END_FUNCTION_BLOCK

// folder: 1000 - 1999 BWT System Control/1130 - 1159 Support Functions

FUNCTION "1130_CALC_TREATMENT_TIME" : LTime   // FC1130, SCL
{ S7_Optimized_Access := 'TRUE' }
VERSION : 0.1
BEGIN
   // Calculate the treatment time of the vessel based on BWMS-066
   #"1130_CALC_TREATMENT_TIME" := "1190_FIXED_CONSTANTS".PreDwell_Time
                                   + ("1190_FIXED_CONSTANTS".DeOxMin_Time * "1191_SYSTEM_VARIABLES".NumberOfActiveTanks)
                                   + "1190_FIXED_CONSTANTS".MidDwell_Time
                                   + "1190_FIXED_CONSTANTS".ReOxMin_Time
                                   + "1190_FIXED_CONSTANTS".PostDwell_Time;
END_FUNCTION

FUNCTION "1131_CALC_HEALTHY_TANKS" : Void   // FC1131, LAD
{ S7_Optimized_Access := 'TRUE' }
VERSION : 0.1
// Calculate which tanks are in a healthy state. If a tank is unhealthy set the deselect flag to True; this will allow the operator the deselect the tank. If the tank is healthy then it must be included in the treatment.
BEGIN

REGION Network 1: If FPT tank is healthy, set deselect to False. (If tank is unhealthy, set Deselect to True)